FUNCTION "Assign_Button.HMI_Stations.WIP" : Void   // FC237, SCL
{ S7_Optimized_Access := 'TRUE' }
VERSION : 0.1
   VAR_INPUT
      processed_inputs : "Settings Screen: Processed Inputs";
      selected_wips : "Selected Wips";
      selected_buttons : "Selected Buttons";
   END_VAR
   VAR_IN_OUT
      pn_library : "Recipe: PN Text Library";
      stations_wips : "WIP: Station";
   END_VAR
   VAR_TEMP
      _i : Int;
      _p_wip : Int;
      _selected_wip_indices : Array[0.."WIP_COUNT"] of Int;
   END_VAR
BEGIN
   REGION "DO NOTHING IF NO WIPS SELECTED"
       IF #selected_wips.count = 0 THEN
           RETURN;
       END_IF;
   END_REGION


   REGION "GET INDICES OF SELECTED WIPS"    
       "WIP_Station.Indices_of_Selected_WIPs"(selected_wips := #selected_wips,
                                              station_wips := #stations_wips,
                                              selected_wip_indices := #_selected_wip_indices);
   END_REGION


   REGION "FOR EACH SELECTED WIP"
       FOR #_i := 0 TO #selected_wips.count DO

           REGION "ASSIGN DATA TO SELECTED BUTTONS"
               #_p_wip := #_selected_wip_indices[#_i];
               IF #_p_wip = "NULL_TOKEN" THEN
                   RETURN;
               END_IF;
               "Assign_Button.HMI_Stations.WIP.Buttons"(processed_inputs := #processed_inputs,
                                                        selected_buttons := #selected_buttons,
                                                        pn_library := #pn_library,
                                                        wip_module := #stations_wips.wip[#_p_wip]);
           END_REGION

       END_FOR;
   END_REGION
END_FUNCTION

FUNCTION "Assign_Button.HMI_Stations.WIP.Buttons" : Void   // FC238, SCL
{ S7_Optimized_Access := 'TRUE' }
VERSION : 0.1
   VAR_INPUT
      processed_inputs : "Settings Screen: Processed Inputs";
      selected_buttons : "Selected Buttons";
   END_VAR
   VAR_IN_OUT
      pn_library : "Recipe: PN Text Library";
      wip_module : "Station: Wip: Wip Module";
   END_VAR
   VAR_TEMP
      _i : Int;
      _p_btn : Int;
      _selected_buttons_indices : Array[0..7] of Int;
   END_VAR
BEGIN
   REGION "DO NOTHING IF NO BUTTONS SELECTED
       IF #selected_buttons.count = 0 THEN
           RETURN;
       END_IF;
   END_REGION


   REGION "GET INDICES OF SELECTED BUTTONS"
       "Selected_Buttons.Indices"(selected_buttons := #selected_buttons,
                                  selected_buttons_indices := #_selected_buttons_indices);
   END_REGION

   REGION "FOR EACH SELECTED BUTTON"
       FOR #_i := 0 TO #selected_buttons.count DO

           REGION "ASSIGN DATA TO SELECTED BUTTON"
               #_p_btn := #_selected_buttons_indices[#_i];
               "Assign_Button.HMI_Stations.Assign_Station_Button_Data"(processed_inputs := #processed_inputs,
                                                                       index := #_p_btn,
                                                                       pn_library := #pn_library,
                                                                       wip_module := #wip_module);
           END_REGION

       END_FOR;
   END_REGION
END_FUNCTION

FUNCTION "Assign_Button.HMI_Stations.Assign_Station_Button_Data" : Void   // FC239, SCL
{ S7_Optimized_Access := 'TRUE' }
VERSION : 0.1
   VAR_INPUT
      processed_inputs : "Settings Screen: Processed Inputs";
      index : Int;
   END_VAR
   VAR_IN_OUT
      pn_library : "Recipe: PN Text Library";
      wip_module : "Station: Wip: Wip Module";
   END_VAR
BEGIN
   IF #index = "NULL_TOKEN" THEN
       RETURN;
   END_IF;
   #wip_module.pnCode[#index] := "Part_Number.WString_to_Code"(part_number := #processed_inputs.part_number.actual,
                                                               pn_library := #pn_library);
   #wip_module.timers.ptAllotted[#index] := #processed_inputs.total.actual;
   #wip_module.timers.ptCritical[#index] := #processed_inputs.critical.actual;
END_FUNCTION

// folder: HMI: Warehouse/002 Settings/Assign Button/KP8 Station

FUNCTION "Assign_Button.KP8_Station" : Void   // FC247, SCL
{ S7_Optimized_Access := 'TRUE' }
VERSION : 0.1
   VAR_INPUT
      processed_inputs : "Settings Screen: Processed Inputs";
      settings : "Settings";
      settings_meta : "Setting Meta Data";
   END_VAR
   VAR_IN_OUT
      all_stations : "Station: All Stations";
      pn_library : "Recipe: PN Text Library";
   END_VAR
   VAR_TEMP
      _i : Int;
      _length : Int;
      _selected_stations : Array[0.."STATION_COUNT"] of Int;
      _p_station : Int;
   END_VAR
BEGIN
   REGION "DO NOTHING IF NO STATIONS SELECTED"
       IF #settings_meta.selected_stations.count = 0 THEN
           RETURN;
       END_IF;
   END_REGION


   REGION "GET INDICES OF SELECTED STATIONS"
       "Selected_Stations.Indices"(selected_stations := #settings_meta.selected_stations,
                                   selected_stations_indices := #_selected_stations);
   END_REGION


   REGION "FOR EACH SELECTED STATION"
       IF #settings_meta.selectable_stations.count = 0 THEN
           RETURN;
       END_IF;
       FOR #_i := 0 TO #settings_meta.selected_stations.count DO
           IF #_selected_stations[#_i] = "NULL_TOKEN" THEN
               RETURN;
           END_IF;
           #_p_station := #_selected_stations[#_i];
           "Assign_Button.Assign_ID_Parameters"(processed_inputs := #processed_inputs,
                                                settings := #settings,
                                                id := #all_stations.stn[#_p_station].id);
           "Assign_Button.KP8_Stations.Buttons"(processed_inputs := #processed_inputs,
                                                selected_buttons := #settings_meta.selected_btns,
                                                pn_library := #pn_library,
                                                station := #all_stations.stn[#_p_station]);
       END_FOR;
   END_REGION
END_FUNCTION

FUNCTION "Assign_Button.KP8_Station.Assign_Station_Button_Data" : Void   // FC248, SCL
{ S7_Optimized_Access := 'TRUE' }
VERSION : 0.1
   VAR_INPUT
      button_number : Int;
      processed_inputs : "Settings Screen: Processed Inputs";
   END_VAR
   VAR_IN_OUT
      pn_library : "Recipe: PN Text Library";
      station : "Station: Single Station";
   END_VAR
   VAR_TEMP
      _i : Int;
      _length : Int;
      _selected_stations : Array[0.."STATION_COUNT"] of Int;
      _p_station : Int;
   END_VAR
BEGIN
   IF #button_number = "NULL_TOKEN" THEN
       RETURN;
   END_IF;
   #station.wipCmpts.pnCode[#button_number] := "Part_Number.WString_to_Code"(part_number := #processed_inputs.part_number.actual,
                                                                             pn_library := #pn_library);
   #station.wipCmpts.timers.ptCritical[#button_number] := #processed_inputs.critical.actual;
   #station.wipCmpts.timers.ptAllotted[#button_number] := #processed_inputs.total.actual;
END_FUNCTION

FUNCTION "Assign_Button.KP8_Stations.Buttons" : Void   // FC249, SCL
{ S7_Optimized_Access := 'TRUE' }
VERSION : 0.1
   VAR_INPUT
      processed_inputs : "Settings Screen: Processed Inputs";
      selected_buttons : "Selected Buttons";
   END_VAR
   VAR_IN_OUT
      pn_library : "Recipe: PN Text Library";
      station : "Station: Single Station";
   END_VAR
   VAR_TEMP
      _i : Int;
      _p_btn : Int;
      _selected_buttons_indices : Array[0..7] of Int;
   END_VAR
BEGIN
   REGION "DO NOTHING IF NO BUTTONS SELECTED
       IF #selected_buttons.count = 0 THEN
           RETURN;
       END_IF;
   END_REGION


   REGION "GET INDICES OF SELECTED BUTTONS"
       "Selected_Buttons.Indices"(selected_buttons := #selected_buttons,
                                  selected_buttons_indices := #_selected_buttons_indices);
   END_REGION


   REGION "FOR EACH SELECTED BUTTON"
       FOR #_i := 0 TO #selected_buttons.count - 1 DO

           IF #_selected_buttons_indices[#_i] = "NULL_TOKEN" THEN
               RETURN;
           END_IF;

           REGION "ASSIGN DATA TO SELECTED BUTTON"
               #_p_btn := #_selected_buttons_indices[#_i];
               "Assign_Button.KP8_Station.Assign_Station_Button_Data"(button_number := #_p_btn,
                                                                      processed_inputs := #processed_inputs,
                                                                      pn_library := #pn_library,
                                                                      station := #station);
           END_REGION

       END_FOR;
   END_REGION
END_FUNCTION

// folder: HMI: Warehouse/002 Settings/Critical IO Field

FUNCTION_BLOCK "Critical_IO_Field"   // FB53, SCL
{ S7_Optimized_Access := 'TRUE' }
VERSION : 0.1
   VAR_INPUT
      settings_meta : "Setting Meta Data";
      stations : "Station: All Stations";
   END_VAR
   VAR_IN_OUT
      interface : "IO Field Data: Label with Data";
      state_changes : "State Changes: Real";
   END_VAR
   VAR
      Critical_IO_Field : "IO Field: State Changes";
      Detect_Stat_Changes : "Real.State_Change";
   END_VAR
   VAR_TEMP
      _interface : "IO Field Data: Label with Data";
      feedback : "IO Field: State Change Data";
   END_VAR
BEGIN
   REGION "BUFFER IN"
       #_interface := #interface;
   END_REGION

   REGION "PROCESS USER INPUT"
       #Critical_IO_Field(interface := #_interface,
                          feedback := #feedback);
       #Detect_Stat_Changes(value := "Timer.WString_to_Real"(#_interface.value),
                            get_real := #state_changes);
   END_REGION

   REGION "BUFFER OUT"
       "Critical_IO_Field.Animate"(feedback := #feedback,
                                   settings_meta := #settings_meta,
                                   stations := #stations,
                                   interface := #_interface);
   END_REGION

   REGION "BUFFER OUT"
       #interface := #_interface;
   END_REGION
END_FUNCTION_BLOCK

FUNCTION "Critical_IO_Field.Make_Visible_Enable" : Bool   // FC191, SCL
{ S7_Optimized_Access := 'TRUE' }
VERSION : 0.1
   VAR_INPUT
      setting_meta : "Setting Meta Data";
   END_VAR
BEGIN
   #"Critical_IO_Field.Make_Visible_Enable" :=  #setting_meta.selected_btns.count > 0;
END_FUNCTION

FUNCTION "Critical_IO_Field.Animate" : Void   // FC192, SCL
{ S7_Optimized_Access := 'TRUE' }
VERSION : 0.1
   VAR_INPUT
      feedback : "IO Field: State Change Data";
      settings_meta : "Setting Meta Data";
      stations : "Station: All Stations";
   END_VAR
   VAR_IN_OUT
      interface : "IO Field Data: Label with Data";
   END_VAR
   VAR_TEMP
      _visible_enabled : Bool;
   END_VAR
BEGIN
   REGION "COLOR"
   #interface.animate := "WHITE_BACKGROUND";
   END_REGION


   REGION "SET STATE"
       #_visible_enabled := "Critical_IO_Field.Make_Visible_Enable"(setting_meta := #settings_meta);
   END_REGION


   REGION "VISIBILITY
       #interface.visible := #_visible_enabled;
   END_REGION


   REGION "ENABLE"
       #interface.enable := #_visible_enabled;
   END_REGION


   REGION "POPULATE VALUE"
       IF #settings_meta.button_selection_change.selection_change THEN
           #interface.value := "Critical_IO_Field.Populate_Value"(hidden := NOT #_visible_enabled,
                                                                  selected_buttons := #settings_meta.selected_btns,
                                                                  selected_stations := #settings_meta.selected_stations,
                                                                  stations := #stations);
       END_IF;
   END_REGION
END_FUNCTION

FUNCTION "Critical_IO_Field.Populate_Value" : WString   // FC283, SCL
{ S7_Optimized_Access := 'TRUE' }
VERSION : 0.1
   VAR_INPUT
      hidden : Bool;
      selected_buttons : "Selected Buttons";
      selected_stations : "Selected Stations";
      stations : "Station: All Stations";
   END_VAR
   VAR_TEMP
      _critical : WString;
      _p_station : Int;
      _p_button : Int;
   END_VAR
   VAR CONSTANT
      BLANK : WString;
      ZERO : WChar := WCHAR#'0';
   END_VAR
BEGIN
   IF #hidden THEN
       #"Critical_IO_Field.Populate_Value" := #BLANK;
       RETURN;
   END_IF;
   #_p_station := "Selected_Stations.Get_First_Selected_Station"(#selected_stations);
   #_p_button := "Selected_Buttons.Get_First_Selected_Button"(#selected_buttons);
   #_critical := "Timer.Real_to_WString"(#stations.stn[#_p_station].wipCmpts.timers.ptCritical[#_p_button]);
   #"Critical_IO_Field.Populate_Value" := #_critical;
END_FUNCTION

// folder: HMI: Warehouse/002 Settings/Dropzone IO Field

FUNCTION_BLOCK "Dropzone_IO_Field"   // FB50, SCL
{ S7_Optimized_Access := 'TRUE' }
VERSION : 0.1
   VAR_INPUT
      settings_meta : "Setting Meta Data";
      stations : "Station: All Stations";
   END_VAR
   VAR_IN_OUT
      interface : "IO Field Data: Label with Data";
      get_dropzone : "State Changes: USInt";
   END_VAR
   VAR
      "Line IO Field" : "IO Field: State Changes";
      "Get Dropzone Input" : "USInt.State_change";
   END_VAR
   VAR_TEMP
      _feedback : "IO Field: State Change Data";
      _interface : "IO Field Data: Label with Data";
   END_VAR
BEGIN
   REGION "BUFFER IN"
       #_interface := #interface;
   END_REGION


   REGION "PROCESS USER INPUT"
       #"Line IO Field"(interface := #_interface,
                        feedback := #_feedback);
       #"Get Dropzone Input"(value := WSTRING_TO_USINT(#interface.value),
                             get_usint := #get_dropzone);
   END_REGION


   REGION "ANIMATION"
       "Dropzone_IO_Field.Animate"(feedback := #_feedback,
                                   selected_stations := #settings_meta.selected_stations,
                                   settings_meta := #settings_meta,
                                   stations := #stations,
                                   interface := #_interface);
   END_REGION


   REGION "BUFFER OUT"
       #interface := #_interface;
   END_REGION
END_FUNCTION_BLOCK

FUNCTION "Dropzone_IO_Field.Make Visible_Enable" : Bool   // FC185, SCL
{ S7_Optimized_Access := 'TRUE' }
VERSION : 0.1
   VAR_INPUT
      setting_meta : "Setting Meta Data";
      stations : "Station: All Stations";
   END_VAR
   VAR_TEMP
      first_selected_station : Int;
      ret : Bool;
   END_VAR
BEGIN
   IF #setting_meta.selected_stations.count = 0 THEN
       #"Dropzone_IO_Field.Make Visible_Enable" := FALSE;
       RETURN;
   END_IF;


   IF #setting_meta.selected_stations.count > 1 THEN
       #"Dropzone_IO_Field.Make Visible_Enable" := FALSE;
       RETURN;
   END_IF;


   IF #setting_meta.selected_btns.count = 0 THEN
       #"Dropzone_IO_Field.Make Visible_Enable"  := FALSE;
       RETURN;
   END_IF;


   #"Dropzone_IO_Field.Make Visible_Enable" := TRUE;
END_FUNCTION

FUNCTION "Dropzone_IO_Field.Animate" : Void   // FC186, SCL
{ S7_Optimized_Access := 'TRUE' }
VERSION : 0.1
   VAR_INPUT
      feedback : "IO Field: State Change Data";
      selected_stations : "Selected Stations";
      settings_meta : "Setting Meta Data";
      stations : "Station: All Stations";
   END_VAR
   VAR_IN_OUT
      interface : "IO Field Data: Label with Data";
   END_VAR
   VAR_TEMP
      _visible_enabled : Bool;
   END_VAR
BEGIN
   REGION "COLOR"
       #interface.animate := "WHITE_BACKGROUND";
   END_REGION


   REGION "GET STATE"
       #_visible_enabled := "Dropzone_IO_Field.Make Visible_Enable"(setting_meta := #settings_meta,
                                                                                stations := #stations);
   END_REGION


   REGION "VISIBILITY
       #interface.visible := #_visible_enabled;
   END_REGION


   REGION "ENABLE"
       #interface.enable := #_visible_enabled;
   END_REGION


   REGION "POPULATE VALUE"
       IF #settings_meta.button_selection_change.selection_change THEN
           #interface.value := "Dropzone_IO_Field.Populate_Value"(hidden := NOT #_visible_enabled,
                                                                  selected_stations := #selected_stations,
                                                                  stations := #stations);
       END_IF;
   END_REGION
END_FUNCTION

FUNCTION "Dropzone_IO_Field.Populate_Value" : WString   // FC271, SCL
{ S7_Optimized_Access := 'TRUE' }
VERSION : 0.1
   VAR_INPUT
      hidden : Bool;
      selected_stations : "Selected Stations";
      stations : "Station: All Stations";
   END_VAR
   VAR_TEMP
      _dropzone : WString;
      _p_station : Int;
   END_VAR
   VAR CONSTANT
      BLANK : WString;
      ZERO : WChar := WCHAR#'0';
   END_VAR
BEGIN
   IF #hidden THEN
       #"Dropzone_IO_Field.Populate_Value" := #BLANK;
       RETURN;
   END_IF;
   #_p_station := "Selected_Stations.Get_First_Selected_Station"(#selected_stations);
   #_dropzone := USINT_TO_WSTRING(#stations.stn[#_p_station].id.dropZone);
   #_dropzone := "Strip Sign"(#_dropzone);
   #_dropzone := "Trim"(#_dropzone);
   #_dropzone := "Add Leading"("Leading Character" := #ZERO,
                               "Desired Length" := 2,
                               "String" := #_dropzone);
   #"Dropzone_IO_Field.Populate_Value" := #_dropzone;
END_FUNCTION

// folder: HMI: Warehouse/002 Settings/Line IO Field

FUNCTION_BLOCK "Line_IO_Field"   // FB47, SCL
{ S7_Optimized_Access := 'TRUE' }
VERSION : 0.1
   VAR_INPUT
      settings_meta : "Setting Meta Data";
      stations : "Station: All Stations";
   END_VAR
   VAR_IN_OUT
      interface : "IO Field Data: Label with Data";
      get_line : "State Changes: WString";
   END_VAR
   VAR
      "Get Line Value" : "WString.State_Change";
      "Line IO Field" : "IO Field: State Changes";
   END_VAR
   VAR_TEMP
      _interface : "IO Field Data: Label with Data";
      feedback : "IO Field: State Change Data";
   END_VAR
BEGIN
   REGION "BUFFER IN"
       #_interface := #interface;
   END_REGION

   REGION "PROCESS USER INPUT"
       #"Line IO Field"(interface := #_interface,
                        feedback := #feedback);
       #"Get Line Value"(interface := #_interface.value,
                         get_wstring := #get_line);

   END_REGION

   REGION "ANIMATION"
       "Line_IO_Field.Animate"(feedback := #feedback,
                               selected_stations := #settings_meta.selected_stations,
                               settings_meta := #settings_meta,
                               stations := #stations,
                               interface := #_interface);
   END_REGION

   REGION "BUFFER OUT"
       #interface := #_interface;
   END_REGION
END_FUNCTION_BLOCK

FUNCTION "Line_IO_Field.Animate" : Void   // FC124, SCL
{ S7_Optimized_Access := 'TRUE' }
VERSION : 0.1
   VAR_INPUT
      feedback : "IO Field: State Change Data";
      selected_stations : "Selected Stations";
      settings_meta : "Setting Meta Data";
      stations : "Station: All Stations";
   END_VAR
   VAR_IN_OUT
      interface : "IO Field Data: Label with Data";
   END_VAR
   VAR_TEMP
      _visible_and_enabled : Bool;
   END_VAR
BEGIN
   REGION "COLOR"
       #interface.animate := "WHITE_BACKGROUND";
   END_REGION


   REGION "STATE"
       #_visible_and_enabled := "Line_IO_Field.Make_Visible_Enable"(selected_stations:= #selected_stations,
                                                                    setting_meta := #settings_meta,
                                                                    stations := #stations);
   END_REGION


   REGION "VISIBILITY
       #interface.visible := #_visible_and_enabled;
   END_REGION


   REGION "ENABLE"
       #interface.enable := #_visible_and_enabled;
   END_REGION


   REGION "POPULATE VALUE"
       IF #settings_meta.button_selection_change.selection_change THEN
           #interface.value := "Line_IO_Field.Populate_Value"(hidden := NOT #_visible_and_enabled,
                                                              selected_stations := #selected_stations,
                                                              stations := #stations);
       END_IF;
   END_REGION
END_FUNCTION

FUNCTION "Line_IO_Field.Make_Visible_Enable" : Bool   // FC187, SCL
{ S7_Optimized_Access := 'TRUE' }
VERSION : 0.1
   VAR_INPUT
      selected_stations : "Selected Stations";
      setting_meta : "Setting Meta Data";
      stations : "Station: All Stations";
   END_VAR
   VAR_TEMP
      first_selected_station : Int;
      ret : Bool;
   END_VAR
BEGIN
   IF #setting_meta.selected_stations.count = 0 THEN
       #"Line_IO_Field.Make_Visible_Enable" := FALSE;
       RETURN;
   END_IF;

   IF #setting_meta.selected_btns.count = 0 THEN
       #"Line_IO_Field.Make_Visible_Enable" := FALSE;
       RETURN;
   END_IF;

   #"Line_IO_Field.Make_Visible_Enable" := "Selected_Stations.Matching_Line_Names"(stations := #stations,
                                                                                               selected_stations := #selected_stations);
END_FUNCTION

FUNCTION "Line_IO_Field.Populate_Value" : WString   // FC268, SCL
{ S7_Optimized_Access := 'TRUE' }
VERSION : 0.1
   VAR_INPUT
      hidden : Bool;
      selected_stations : "Selected Stations";
      stations : "Station: All Stations";
   END_VAR
   VAR_TEMP
      _p_station : Int;
   END_VAR
   VAR CONSTANT
      BLANK : WString;
   END_VAR
BEGIN
   IF #hidden THEN
       #"Line_IO_Field.Populate_Value" := #BLANK;
       RETURN;
   END_IF;
   #_p_station := "Selected_Stations.Get_First_Selected_Station"(#selected_stations);
   #"Line_IO_Field.Populate_Value" := #stations.stn[#_p_station].id.lineName;
END_FUNCTION

// folder: HMI: Warehouse/002 Settings/Part Number IO Field

FUNCTION_BLOCK "Part Number IO Field"   // FB54, SCL
{ S7_Optimized_Access := 'TRUE' }
VERSION : 0.1
   VAR_INPUT
      settings_meta : "Setting Meta Data";
      stations : "Station: All Stations";
      part_number_library : "Recipe: PN Text Library";
   END_VAR
   VAR_IN_OUT
      interface : "Part_Number_Double.UDT";
      processed_part_number_entry : "State Changes: WString";
   END_VAR
   VAR
      Resolve_Feedback : "Part_Number_Double.State_Changes";
      Get_Part_Number : "Part_Number_IO_Field.Get_Part_Number";
      display_mode : String[10] := 'single';
   END_VAR
   VAR_TEMP
      _interface : "Part_Number_Double.UDT";
      feedback : "Part_Number_Double.State_Change.UDT";
   END_VAR
BEGIN
   REGION "BUFFER IN"
       #_interface := #interface;
   END_REGION


   REGION "PROCESS USER INPUT"
       #Resolve_Feedback(interface := #_interface,
                         feedback := #feedback);
       "Part_Number_Double_IO_Field.Set_Mode"(feedback := #feedback,
                                              mode := #display_mode);
       #Get_Part_Number(mode := #display_mode,
                        feedback := #feedback,
                        processed_part_number_entry := #processed_part_number_entry);
   END_REGION


   REGION "ANIMATE"
       "Part_Number_IO_Field.Animate"(display_mode := #display_mode,
                                      settings_meta := #settings_meta,
                                      stations := #stations,
                                      part_number_library := #part_number_library,
                                      interface := #_interface);
   END_REGION


   REGION "BUFFER OUT"
       #interface := #_interface;
   END_REGION
END_FUNCTION_BLOCK

FUNCTION "Part_Number_IO_Field.Make_Visible_Enable" : Bool   // FC195, SCL
{ S7_Optimized_Access := 'TRUE' }
VERSION : 0.1
   VAR_INPUT
      setting_meta : "Setting Meta Data";
      visible_mode : String;
      current_mode : String;
   END_VAR
BEGIN
   IF #setting_meta.selected_btns.count = 0 THEN
       #"Part_Number_IO_Field.Make_Visible_Enable" := FALSE;
       RETURN;
   END_IF;

   #"Part_Number_IO_Field.Make_Visible_Enable" := #visible_mode = #current_mode;
END_FUNCTION

FUNCTION "Part_Number_IO_Field.Animate" : Void   // FC196, SCL
{ S7_Optimized_Access := 'TRUE' }
VERSION : 0.1
   VAR_INPUT
      settings_meta : "Setting Meta Data";
      stations : "Station: All Stations";
      part_number_library : "Recipe: PN Text Library";
   END_VAR
   VAR_IN_OUT
      display_mode : String;
      interface : "Part_Number_Double.UDT";
   END_VAR
   VAR_TEMP
      _double_visible_enabled : Bool;
      _single_visible_enabled : Bool;
   END_VAR
   VAR CONSTANT
      SINGLE : String := 'single';
      DOUBLE : String := 'double';
   END_VAR
BEGIN
   REGION "COLOR"
       #interface.single_animate := "WHITE_BACKGROUND";
       #interface.double_animate := "WHITE_BACKGROUND";
   END_REGION


   REGION "STATE"
       #_single_visible_enabled := "Part_Number_IO_Field.Make_Visible_Enable"(setting_meta := #settings_meta,
                                                                              visible_mode := #SINGLE,
                                                                              current_mode := #display_mode);
       #_double_visible_enabled := "Part_Number_IO_Field.Make_Visible_Enable"(setting_meta := #settings_meta,
                                                                              visible_mode := #DOUBLE,
                                                                              current_mode := #display_mode);
   END_REGION


   REGION "VISIBILITY"
       #interface.single_visible := #_single_visible_enabled;
       #interface.double_visible := #_double_visible_enabled;
   END_REGION


   REGION "ENABLE"
       #interface.single_enable := #interface.single_visible;
       #interface.double_enable := #interface.double_visible;
   END_REGION


   REGION "POPULATE VALUE"
       IF #settings_meta.button_selection_change.selection_change THEN
           "Part_Number_IO_Field.Populate_Value"(stations := #stations,
                                                 settings_meta := #settings_meta,
                                                 part_number_library := #part_number_library,
                                                 display_mode := #display_mode,
                                                 interface := #interface);
       END_IF;
   END_REGION
END_FUNCTION

FUNCTION "Part_Number_IO_Field.Populate_Value" : Void   // FC293, SCL
{ S7_Optimized_Access := 'TRUE' }
VERSION : 0.1
   VAR_INPUT
      part_number_library : "Recipe: PN Text Library";
      stations : "Station: All Stations";
      settings_meta : "Setting Meta Data";
   END_VAR
   VAR_IN_OUT
      display_mode : String;
      interface : "Part_Number_Double.UDT";
   END_VAR
   VAR_TEMP
      _p_button : Int;
      _p_station : Int;
      _part_number_code : DInt;
      _part_number : WString;
      _split_part_numbers : Array[0..1] of WString;
   END_VAR
   VAR CONSTANT
      SINGLE : String := 'single';
      DOUBLE : String := 'double';
   END_VAR
BEGIN
   #_p_button := "Selected_Buttons.Get_First_Selected_Button"(#settings_meta.selected_btns);
   IF #_p_button = "NULL_TOKEN" THEN
       RETURN;
   END_IF;
   #_p_station := "Selected_Stations.Get_First_Selected_Station"(#settings_meta.selected_stations);
   IF #_p_station = "NULL_TOKEN" THEN
       RETURN;
   END_IF;
   #_part_number_code := #stations.stn[#_p_station].wipCmpts.pnCode[#_p_button];
   #_part_number := "Part_Number.Code_to_WString"(pnLib := #part_number_library,
                                                  pnCode := #_part_number_code);
   IF "Part_Number.Is_Single"(#_part_number_code) THEN
       #interface.single_value := #_part_number;
       #display_mode := #SINGLE;
       RETURN;
   END_IF;
   "Part_Number.Split_PNs"(part_number := #_part_number,
                           part_numbers := #_split_part_numbers);
   #interface.double_value_top := #_split_part_numbers[0];
   #interface.double_value_bottom := #_split_part_numbers[1];
   #display_mode := #DOUBLE;
   RETURN;
END_FUNCTION

// folder: HMI: Warehouse/002 Settings/Select Buttons Button

FUNCTION_BLOCK "Select Buttons"   // FB42, SCL
{ S7_Optimized_Access := 'TRUE' }
VERSION : 0.1
   VAR_INPUT
      settings_meta : "Setting Meta Data";
      stations : "Station: All Stations";
   END_VAR
   VAR_IN_OUT
      interface : "Push Button Data";
   END_VAR
   VAR
      "Get Button Feedback" : "Push Button: State Changes";
   END_VAR
   VAR_TEMP
      _interface : "Push Button Data";
      enable : Bool;
      feedback : "Push Button Data: State Change Data";
      visible : Bool;
   END_VAR
BEGIN
   REGION "BUFFER IN"
       #_interface := #interface;
   END_REGION

   REGION "PROCESS USER INPUT"
       #"Get Button Feedback"(interface := #_interface,
                              state_changes := #feedback);
   END_REGION

   REGION "ANIMATIONS"
       "Select Buttons: Private: Animations"(feedback := #feedback,
                                             settings_meta := #settings_meta,
                                             stations := #stations,
                                             interface := #_interface);
   END_REGION

   REGION "BUFFER OUT"
       #interface := #_interface;
   END_REGION
END_FUNCTION_BLOCK

FUNCTION "Select Buttons: Private: Animations" : Void   // FC93, SCL
{ S7_Optimized_Access := 'TRUE' }
VERSION : 0.1
   VAR_INPUT
      feedback : "Push Button Data: State Change Data";
      settings_meta : "Setting Meta Data";
      stations : "Station: All Stations";
   END_VAR
   VAR_IN_OUT
      interface : "Push Button Data";
   END_VAR
BEGIN
   REGION "COLOR"
       #interface.animate := "Bool.Animate"(true_color := "GREEN_LIGHT_BACKGROUND",
                                             false_color := "GRAY_BACKGROUND",
                                             evaluation_signal := #feedback.actuate.actual);
   END_REGION

   REGION "VISIBILITY"
       #interface.visible := "Select Buttons: Private: Make Visible / Enable"(settings_meta := #settings_meta,
                                                                               stations := #stations);
   END_REGION

   REGION "ENABLED STATE"
       #interface.enable := "Select Buttons: Private: Make Visible / Enable"(settings_meta := #settings_meta,
                                                                              stations := #stations);
   END_REGION
END_FUNCTION

FUNCTION "Select Buttons: Private: Make Visible / Enable" : Bool   // FC184, SCL
{ S7_Optimized_Access := 'TRUE' }
VERSION : 0.1
   VAR_INPUT
      settings_meta : "Setting Meta Data";
      stations : "Station: All Stations";
   END_VAR
   VAR_TEMP
      ret : Bool;
      enable : Bool;
      is_hmi_station : Bool;
   END_VAR
BEGIN
   REGION "STATIONS ARE HMI STATIONS"
       #is_hmi_station := "Is_HMI_Station"(#stations.stn["Get First Selected Station"(#settings_meta.selected_stations.stns)]);
   END_REGION

   REGION "ENABLE/MAKE VISIBLE"
       IF (#settings_meta.selected_stations.count > 0) AND
           ((#is_hmi_station AND #settings_meta.selected_wips.count> 0) OR NOT #is_hmi_station) THEN
               #ret := TRUE;
       END_IF;
   END_REGION

   REGION "RETURN"
       #"Select Buttons: Private: Make Visible / Enable" := #ret;
   END_REGION
END_FUNCTION

// folder: HMI: Warehouse/002 Settings/Select Station Button

FUNCTION_BLOCK "Select Station PB"   // FB45, SCL
{ S7_Optimized_Access := 'TRUE' }
VERSION : 0.1
   VAR_IN_OUT
      interface : "Push Button Data";
   END_VAR
   VAR
      "Get Button Feedback" : "Push Button: State Changes";
   END_VAR
   VAR_TEMP
      _interface : "Push Button Data";
      feedback : "Push Button Data: State Change Data";
   END_VAR
BEGIN
   REGION "BUFFER IN"
       #_interface := #interface;
   END_REGION

   REGION "PROCESS USER INPUT"
       #"Get Button Feedback"(interface := #_interface,
                              state_changes := #feedback);
   END_REGION

   REGION "ANIMATIONS"
       "Select Station PB: Private: Animations"(feedback := #feedback,
                                                interface := #_interface);
   END_REGION

   REGION "BUFFER OUT"
       #interface := #_interface;
   END_REGION
END_FUNCTION_BLOCK

FUNCTION "Select Station PB: Private: Animations" : Void   // FC94, SCL
{ S7_Optimized_Access := 'TRUE' }
VERSION : 0.1
   VAR_INPUT
      feedback : "Push Button Data: State Change Data";
   END_VAR
   VAR_IN_OUT
      interface : "Push Button Data";
   END_VAR
BEGIN
   REGION "COLOR"
       #interface.animate := "Bool.Animate"(true_color := "GREEN_LIGHT_BACKGROUND",
                                             false_color := "GRAY_BACKGROUND",
                                             evaluation_signal := #feedback.actuate.actual);
   END_REGION

   REGION "VISIBILITY"
       #interface.visible := TRUE;
   END_REGION

   REGION "ENABLED STATE"
       #interface.enable := TRUE;
   END_REGION
END_FUNCTION

// folder: HMI: Warehouse/002 Settings/Select WIP Button

FUNCTION_BLOCK "Select WIP PB"   // FB46, SCL
{ S7_Optimized_Access := 'TRUE' }
VERSION : 0.1
   VAR_INPUT
      settings_meta : "Setting Meta Data";
      stations : "Station: All Stations";
   END_VAR
   VAR_IN_OUT
      interface : "Push Button Data";
   END_VAR
   VAR
      "Get Button Feedback" : "Push Button: State Changes";
   END_VAR
   VAR_TEMP
      _interface : "Push Button Data";
      enable : Bool;
      feedback : "Push Button Data: State Change Data";
      visible : Bool;
   END_VAR
BEGIN
   REGION "BUFFER IN"
       #_interface := #interface;
   END_REGION

   REGION "PROCESS USER INPUT"
       #"Get Button Feedback"(interface := #_interface,
                              state_changes := #feedback);
   END_REGION

   REGION "ANIMATIONS"
       "Select WIP PB: Private: Animations"(feedback := #feedback,
                                            settings_meta := #settings_meta,
                                            stations := #stations,
                                            interface := #_interface);
   END_REGION

   REGION "BUFFER OUT"
       #interface := #_interface;
   END_REGION
END_FUNCTION_BLOCK

FUNCTION "Select WIP PB: Private: Make Visible / Enable" : Bool   // FC92, SCL
{ S7_Optimized_Access := 'TRUE' }
VERSION : 0.1
   VAR_INPUT
      settings_meta : "Setting Meta Data";
      stations : "Station: All Stations";
   END_VAR
   VAR_TEMP
      ret : Bool;
      index_of_first_selected_station : Int;
      is_hmi_station : Bool;
      first_selected_station : "Station: Single Station";
      t_select_wip : "Push Button Data";
   END_VAR
BEGIN
   REGION "ARE SELECTED STATIONS HMI STATIONS?"
       #index_of_first_selected_station := "Get First Selected Station"(#settings_meta.selected_stations.stns);
       #first_selected_station := #stations.stn[#index_of_first_selected_station];
       #is_hmi_station := "Is_HMI_Station"(#first_selected_station);
   END_REGION

   REGION "HMI STATIONS"
       IF #is_hmi_station THEN
           #ret := TRUE;
       END_IF;
   END_REGION

   REGION "RETURN"
       #"Select WIP PB: Private: Make Visible / Enable" := #ret;
   END_REGION
END_FUNCTION

FUNCTION "Select WIP PB: Private: Animations" : Void   // FC123, SCL
{ S7_Optimized_Access := 'TRUE' }
VERSION : 0.1
   VAR_INPUT
      feedback : "Push Button Data: State Change Data";
      settings_meta : "Setting Meta Data";
      stations : "Station: All Stations";
   END_VAR
   VAR_IN_OUT
      interface : "Push Button Data";
   END_VAR
BEGIN
   REGION "COLOR"
       #interface.animate := "Bool.Animate"(true_color := "GREEN_LIGHT_BACKGROUND",
                                             false_color := "GRAY_BACKGROUND",
                                             evaluation_signal := #feedback.actuate.actual);
   END_REGION

   REGION "VISIBILITY"
       #interface.visible := "Select WIP PB: Private: Make Visible / Enable"(settings_meta := #settings_meta,
                                                                              stations := #stations);
   END_REGION

   REGION "ENABLED STATE"
       #interface.enable := "Select WIP PB: Private: Make Visible / Enable"(settings_meta := #settings_meta,
                                                                             stations := #stations);
   END_REGION
END_FUNCTION

// folder: HMI: Warehouse/002 Settings/Selected WIP Table

FUNCTION_BLOCK "Selected_WIP_Table"   // FB30, SCL
{ S7_Optimized_Access := 'TRUE' }
VERSION : 0.1
   VAR_INPUT
      navigation_bar : "Nav Bar Data: PLC";
      pn_library : "Recipe: PN Text Library";
      saved_wips : "Recipe: HMI Stations Saved Wips";
      settings_meta : "Setting Meta Data";
      stations : "Station: All Stations";
      wip_library : "Recipe: Wip Text Library";
   END_VAR
   VAR_IN_OUT
      stationRows : Array[0..2] of "Settings Station Row Data";
   END_VAR
   VAR
      first_selected_station : Int;
      hmi_stations_selected : Bool;
      selected_stations : Array[0.."STATION_COUNT"] of Int;
      selected_list : "Selected_WIP_Table.Selected_Array";
      row_indices : Array[0..2] of DInt;
      inst_Table_Navigation : "Table Nav";
   END_VAR
   VAR_TEMP
      i : Int;
      p_stn : Int;
      wip_code : DInt;
      visible_rows : Int;
      first_null_index : DInt;
      _hmi_saved_station_index : Int;
      _wip_index : Int;
      _wip_module : "Station: Wip: Wip Module";
   END_VAR
   // row_indices[0] := 0;
   // row_indices[1] := 1;
   // row_indices[2] := 2;
BEGIN
   REGION "CLEAR OLD CONTENTS"    
       FOR #i := 0 TO 2 DO
           #stationRows[#i].line := "Cell_Data.Hide"();
           #stationRows[#i].dropzone := "Cell_Data.Hide"();
           #stationRows[#i].wip := "Cell_Data.Hide"();
           "Button_Row.Hide_Rows"(#stationRows[#i].btnRows);
       END_FOR;
   END_REGION


   REGION "EXIT ON NO SELECTED STATION"
       IF #settings_meta.selected_stations.count = 0 THEN
           RETURN;
       END_IF;
   END_REGION


   REGION "GET ARRAY OF SELECTED STATION INDICES"
       "Array.Int.Fill"(value := "NULL_TOKEN",
                        int_array := #selected_stations);
       "Selected_Stations.Indices"(selected_stations := #settings_meta.selected_stations,
                                   selected_stations_indices := #selected_stations);
       "Selected_WIP_Table.Build_List"(selected_stations := #selected_stations,
                                       selected_wips := #settings_meta.selected_wips.wips,
                                       selected_list := #selected_list);
   END_REGION


   REGION "DETERMINE IF SELECTED STATION IS AN HMI STATION"
       #first_selected_station := "Get First Selected Station"(#settings_meta.selected_stations.stns);
       #hmi_stations_selected := "Is_HMI_Station"(#stations.stn[#first_selected_station]);
   END_REGION


   REGION "TABLE DISPLAY POINTERS"
       #first_null_index := "Selected_WIP_Table.Selected_Array.First_Occurance"(selected_array := #selected_list,
                                                                                search_term := "NULL_TOKEN");
       #inst_Table_Navigation(first_null_index := #first_null_index,
                              tblData := #selected_list.me,
                              tblDisp := #stationRows,
                              tableNav := #navigation_bar,
                              rowIndices := #row_indices);
   END_REGION


   REGION "TABLE COMPONENTS"
       #visible_rows := DINT_TO_INT(#first_null_index) - 1;
       IF #visible_rows > 2 THEN
           #visible_rows := 2;
       END_IF;
       FOR #i := 0 TO #visible_rows DO
           #p_stn := #selected_list.me[#row_indices[#i]].station_pointer;
           #wip_code := #selected_list.me[#row_indices[#i]].wip_pointer;
           #stationRows[#i].line := "Selected_WIP_Table.Line_Label.Show"(station := #stations.stn[#p_stn]);
           #stationRows[#i].dropzone := "Selected_WIP_Table.Dropzone_Label.Show"(station := #stations.stn[#p_stn]);
           #stationRows[#i].wip := "Selected_WIP_Table.Wip_Label.Show"(wip_code := #wip_code,
                                                                       wip_library := #wip_library);
           #_wip_module := "Selected_WIP_Table.Get_WIP_Module"(stations := #stations,
                                                               saved_wips := #saved_wips,
                                                               station_pointer := #p_stn,
                                                               wip_code := #wip_code);
           "Button_Row.Show_Rows"(selected_butttons := #settings_meta.selected_btns,
                                  wip_module := #_wip_module,
                                  pn_library := #pn_library,
                                  button_rows := #stationRows[#i].btnRows);
       END_FOR;
   END_REGION
END_FUNCTION_BLOCK

FUNCTION "Selected_WIP_Table.Build_List" : Void   // FC219, SCL
{ S7_Optimized_Access := 'TRUE' }
VERSION : 0.1
   VAR_INPUT
      selected_stations : Array[*] of Int;
      selected_wips : Array[*] of DInt;
   END_VAR
   VAR_IN_OUT
      selected_list : "Selected_WIP_Table.Selected_Array";
   END_VAR
   VAR_TEMP
      _i : DInt;
      _j : DInt;
      _length : Struct
         stations : DInt;
         wips : DInt;
      END_STRUCT;
      _p : DInt;
   END_VAR
BEGIN
   REGION "PREPARE ARRAY"
       "Selected_WIP_Table.Selected_Array.Fill"(token := -1,
                                                selected_list := #selected_list);
   END_REGION


   REGION "GET UPPER LIMIT FOR OUTER LOOP"
       #_length.stations := "Array.Int.First_Occurance"(int_array := #selected_stations,
                                                        search_term := "NULL_TOKEN");
       #_length.stations -= 1;
       #_length.stations := "DInt.Clip.Minimum"(value := #_length.stations,
                                                minimum := 0);
   END_REGION


   REGION "GET LIMIT FOR INNER LOOP"
       #_length.wips := "Array.DInt.First_Occurance"(dint_array := #selected_wips,
                                                     search_term := "NULL_TOKEN");
       #_length.wips -= 1;
       #_length.wips := "DInt.Clip.Minimum"(value := #_length.wips,
                                            minimum := 0);
   END_REGION


   REGION "BUILD ARRAY"
       FOR #_i := 0 TO #_length.stations DO
           FOR #_j := 0 TO #_length.wips DO
               #_p := #_i * (#_length.wips + 1) + #_j;
               #selected_list.me[#_p].station_pointer := #selected_stations[#_i];
               #selected_list.me[#_p].wip_pointer := #selected_wips[#_j];
           END_FOR;
       END_FOR;
   END_REGION
END_FUNCTION

FUNCTION "Selected_WIP_Table.Selected_Array.Fill" : Void   // FC221, SCL
{ S7_Optimized_Access := 'TRUE' }
VERSION : 0.1
   VAR_INPUT
      token : Int;
   END_VAR
   VAR_IN_OUT
      selected_list : "Selected_WIP_Table.Selected_Array";
   END_VAR
   VAR_TEMP
      _i : DInt;
      _length : DInt;
   END_VAR
BEGIN
   #_length := UDINT_TO_DINT("Array.Any.Length"(#selected_list.me));
   #_length -= 1;

   FOR #_i := 0 TO #_length DO
       #selected_list.me[#_i].station_pointer := #token;
       #selected_list.me[#_i].wip_pointer := INT_TO_DINT(#token);
   END_FOR;
END_FUNCTION

FUNCTION "Selected_WIP_Table.Selected_Array.Is_Element" : Bool   // FC228, SCL
{ S7_Optimized_Access := 'TRUE' }
VERSION : 0.1
   VAR_INPUT
      selected_array : "Selected_WIP_Table.Selected_Array";
      search_term : Int;
   END_VAR
   VAR_TEMP
      _i : DInt;
      _length : DInt;
   END_VAR
BEGIN
   REGION "LOCAL VARIABLES"
       #_length := UDINT_TO_DINT("Array.Any.Length"(#selected_array.me)) - 1;
   END_REGION


   REGION "SEARCH ARRAY"
       FOR #_i := 0 TO #_length DO
           IF #selected_array.me[#_i].station_pointer <> #search_term THEN
               CONTINUE;
           END_IF;
           #"Selected_WIP_Table.Selected_Array.Is_Element" := TRUE;
           RETURN;
       END_FOR;
   END_REGION


   REGION "NOT FOUND"
       #"Selected_WIP_Table.Selected_Array.Is_Element" := FALSE;
       RETURN;
   END_REGION
END_FUNCTION

FUNCTION "Selected_WIP_Table.Selected_Array.First_Occurance" : DInt   // FC229, SCL
{ S7_Optimized_Access := 'TRUE' }
VERSION : 0.1
   VAR_INPUT
      selected_array : "Selected_WIP_Table.Selected_Array";
      search_term : Int;
   END_VAR
   VAR_TEMP
      _i : DInt;
      _length : UDInt;
   END_VAR
BEGIN
   REGION "NOTES"
       (* 
       This function returns the first occurance of the search term.
       This function meant for use with collapsed arrays.
       See "Array.Int.Collapse" for collapse functionality.
       *)
   END_REGION


   REGION "GET LENGTH OF INPUT ARRAY"
       #_length := "Array.Any.Length"(#selected_array.me);
   END_REGION


   REGION "FIND FIRST SEARCH TERM, -1 IF NONE"
       (*
       Its worth noting that "Array.Int.Is_Element" could return the index of the search term
       as an output, saving the processor some work. 
       The rework is justified by increased encapsulation.
       The time complexity for "Array.Int.First_Occurance" remains O(n).
       *)
       IF NOT "Selected_WIP_Table.Selected_Array.Is_Element"(selected_array:=#selected_array, search_term:=#search_term) THEN
           #"Selected_WIP_Table.Selected_Array.First_Occurance" := -1;
           RETURN;
       END_IF;
       WHILE #selected_array.me[#_i].station_pointer <> #search_term AND DINT_TO_UDINT(#_i) < #_length DO
           #_i += 1;
       END_WHILE;
   END_REGION


   REGION "SEARCH TERM FOUND"
       #"Selected_WIP_Table.Selected_Array.First_Occurance" := #_i;
       RETURN;
   END_REGION
END_FUNCTION

FUNCTION "Selected_WIP_Table.Get_WIP_Module" : "Station: Wip: Wip Module"   // FC234, SCL
{ S7_Optimized_Access := 'TRUE' }
VERSION : 0.1
   VAR_INPUT
      stations : "Station: All Stations";
      saved_wips : "Recipe: HMI Stations Saved Wips";
      station_pointer : Int;
      wip_code : DInt;
   END_VAR
   VAR_TEMP
      _hmi_station_pointer : Int;
      _wip_pointer : Int;
   END_VAR
BEGIN
   IF #wip_code = "NULL_TOKEN" THEN
       #"Selected_WIP_Table.Get_WIP_Module" := #stations.stn[#station_pointer].wipCmpts;
       RETURN;
   END_IF;

   #_hmi_station_pointer := "WIP.Global_Index_to_HMI_Station_Index"(global_index := #station_pointer,
                                                                    saved_WIPs := #saved_wips);

   #_wip_pointer := "WIP.Code_to_Index"(saved_wip := #saved_wips.stn[#_hmi_station_pointer],
                                        wip_code := #wip_code);

   #"Selected_WIP_Table.Get_WIP_Module" := #saved_wips.stn[#_hmi_station_pointer].wip[#_wip_pointer];
   RETURN;
END_FUNCTION

// folder: HMI: Warehouse/002 Settings/Selected WIP Table/Button Row

FUNCTION "Button_Row.Hide" : "Settings Station Row Button Row Data"   // FC210, SCL
{ S7_Optimized_Access := 'TRUE' }
VERSION : 0.1
   VAR_TEMP
      _ret : "Settings Station Row Button Row Data";
   END_VAR
BEGIN
   #_ret.button := "Cell_Data.Hide"();
   #_ret.total := "Cell_Data.Hide"();
   #_ret.critical := "Cell_Data.Hide"();
   #_ret.singlePN := "Cell_Data.Hide"();
   #_ret.doublePN := "Cell_Data.Hide"();
   #"Button_Row.Hide" := #_ret;
END_FUNCTION

FUNCTION "Button_Row.Hide_Rows" : Void   // FC211, SCL
{ S7_Optimized_Access := 'TRUE' }
VERSION : 0.1
   VAR_IN_OUT
      button_rows : Array[*] of "Settings Station Row Button Row Data";
   END_VAR
   VAR_TEMP
      _i : Int;
   END_VAR
BEGIN
   FOR #_i := 0 TO UDINT_TO_INT("Array.Any.Length"(#button_rows)) - 1 DO
       #button_rows[#_i] := "Button_Row.Hide"();
   END_FOR;
END_FUNCTION

FUNCTION "Button_Row.Show" : "Settings Station Row Button Row Data"   // FC212, SCL
{ S7_Optimized_Access := 'TRUE' }
VERSION : 0.1
   VAR_INPUT
      button_number : Int;
      selected : Bool;
      pn_library : "Recipe: PN Text Library";
      wip_module : "Station: Wip: Wip Module";
   END_VAR
   VAR_TEMP
      _return : "Settings Station Row Button Row Data";
      _pn : "Cell Data";
   END_VAR
BEGIN
   #_return.button := "Button_Row.Button_Label.Show"(button_number := #button_number,
                                                     selected := #selected);

   #_return.total := "Button_Row.Total.Show"(selected := #selected,
                                             button_number := #button_number,
                                             wip_module := #wip_module);

   #_return.critical := "Button_Row.Critical.Show"(button_number := #button_number,
                                                   selected := #selected,
                                                   wip_module := #wip_module);

   #_pn := "Button_Row.Part_Number.Show"(button_number := #button_number,
                                         pn_library := #pn_library,
                                         selected := #selected,
                                         wip_module := #wip_module);

   IF "Part_Number.Is_Single"(#wip_module.pnCode[#button_number]) THEN
       #_return.singlePN := #_pn;
   END_IF;
   IF "Part_Number.Is_Double"(#wip_module.pnCode[#button_number]) THEN
       #_return.doublePN := #_pn;
   END_IF;
   #"Button_Row.Show" := #_return;
END_FUNCTION

FUNCTION "Button_Row.Show_Rows" : Void   // FC218, SCL
{ S7_Optimized_Access := 'TRUE' }
VERSION : 0.1
   VAR_INPUT
      selected_butttons : "Selected Buttons";
      wip_module : "Station: Wip: Wip Module";
      pn_library : "Recipe: PN Text Library";
   END_VAR
   VAR_IN_OUT
      button_rows : Array[*] of "Settings Station Row Button Row Data";
   END_VAR
   VAR_TEMP
      _i : Int;
      _remap : Int;
   END_VAR
BEGIN
   FOR #_i := 0 TO UDINT_TO_INT("Array.Any.Length"(#button_rows)) - 1 DO
       #_remap := "KP8.DURL_to_LRUD"(#_i);
       #button_rows[#_i] := "Button_Row.Show"(button_number := #_remap,
                                              selected := #selected_butttons.btns[#_i],
                                              pn_library := #pn_library,
                                              wip_module := #wip_module);
   END_FOR;
END_FUNCTION

// folder: HMI: Warehouse/002 Settings/Selected WIP Table/Button Row/Single Button